REGION Network 13
   "V003 - Ventilador 3 Torres de enfriamiento Chillers"(Input_0 := "V003-TO",   // "FB_CTR_MOT"
                           Input_1 := "V003-CO",
                           Input_3 := ("DB90".Static_142 OR ("DB92".Static_12 AND NOT "DB90".Static_12)) AND NOT "DB86".Static_67 AND NOT "DB86".Static_68,
                           Input_6 := "UNO",
                           Input_7 := "DB90".Static_116,
                           Input_8 := "DB90".Static_12,
                           Output_0 => "V003-Marcha",
                           Output_2 => "DB32".Static_35,
                           Output_3 => "DB32".Static_36);
END_REGION

REGION Network 14
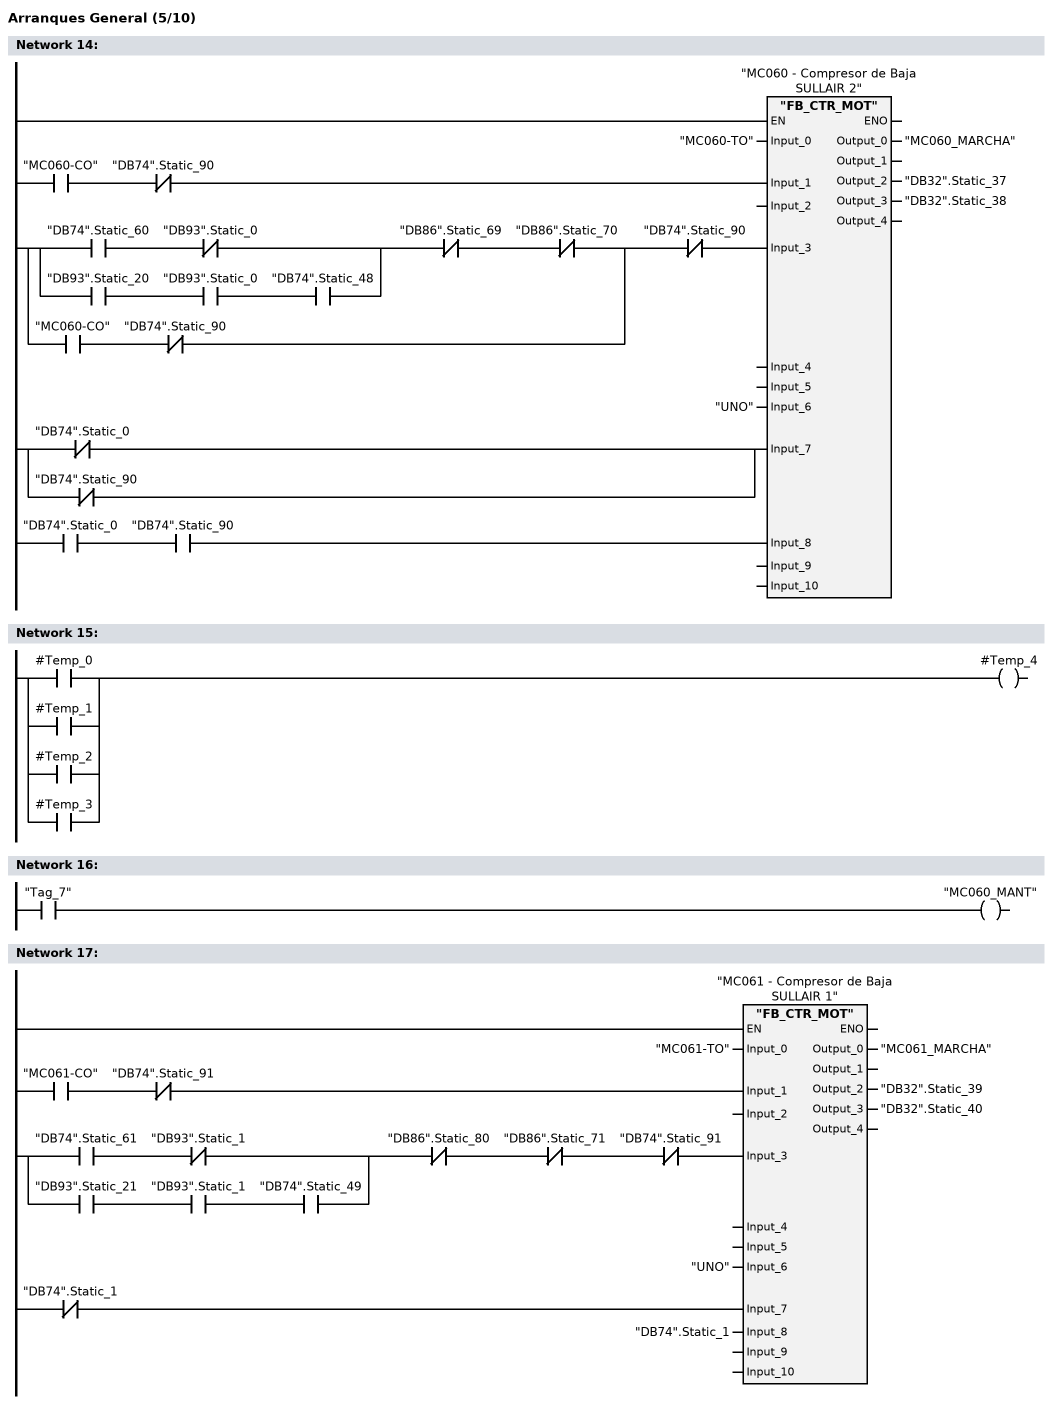
   "MC060 - Compresor de Baja SULLAIR 2"(Input_0 := "MC060-TO",   // "FB_CTR_MOT"
                           Input_1 := "MC060-CO" AND NOT "DB74".Static_90,
                           Input_3 := (((("DB74".Static_60 AND NOT "DB93".Static_0) OR ("DB93".Static_20 AND "DB93".Static_0 AND "DB74".Static_48)) AND NOT "DB86".Static_69 AND NOT "DB86".Static_70) OR ("MC060-CO" AND NOT "DB74".Static_90)) AND NOT "DB74".Static_90,
                           Input_6 := "UNO",
                           Input_7 := NOT "DB74".Static_0 OR NOT "DB74".Static_90,
                           Input_8 := "DB74".Static_0 AND "DB74".Static_90,
                           Output_0 => "MC060_MARCHA",
                           Output_2 => "DB32".Static_37,
                           Output_3 => "DB32".Static_38);
END_REGION

REGION Network 15
   RUNG wire#powerrail
      Contact( #Temp_0 )
      wire#w1
      Coil( #Temp_4 )
   END_RUNG
   RUNG wire#powerrail
      Contact( #Temp_1 )
   END_RUNG wire#w1
   RUNG wire#powerrail
      Contact( #Temp_2 )
   END_RUNG wire#w1
   RUNG wire#powerrail
      Contact( #Temp_3 )
   END_RUNG wire#w1
   // the same network as SCL:
   #Temp_4 := #Temp_0 OR #Temp_1 OR #Temp_2 OR #Temp_3;
END_REGION

REGION Network 16
   RUNG wire#powerrail
      Contact( "Tag_7" )
      Coil( "MC060_MANT" )
   END_RUNG
   // the same network as SCL:
   "MC060_MANT" := "Tag_7";
END_REGION

REGION Network 17
   RUNG wire#powerrail
      "MC061 - Compresor de Baja SULLAIR 1"(Input_0 := "MC061-TO", Input_2 :=, Input_4 :=, Input_5 :=, Input_6 := "UNO", Input_8 := "DB74".Static_1, Input_9 :=, Input_10 :=, Output_0 => "MC061_MARCHA", Output_1 =>, Output_2 => "DB32".Static_39, Output_3 => "DB32".Static_40, Output_4 =>, Input_1 := wire#w1, Input_3 := wire#w3, Input_7 := wire#w4)
   END_RUNG
   RUNG wire#powerrail
      Contact( "MC061-CO" )
      I_Contact( "DB74".Static_91 )
   END_RUNG wire#w1
   RUNG wire#powerrail
      Contact( "DB74".Static_61 )
      I_Contact( "DB93".Static_1 )
      wire#w2
      I_Contact( "DB86".Static_80 )
      I_Contact( "DB86".Static_71 )
      I_Contact( "DB74".Static_91 )
   END_RUNG wire#w3
   RUNG wire#powerrail
      Contact( "DB93".Static_21 )
      Contact( "DB93".Static_1 )
      Contact( "DB74".Static_49 )
   END_RUNG wire#w2
   RUNG wire#powerrail
      I_Contact( "DB74".Static_1 )
   END_RUNG wire#w4
   // the same network as SCL:
   "MC061 - Compresor de Baja SULLAIR 1"(Input_0 := "MC061-TO",   // "FB_CTR_MOT"
                           Input_1 := "MC061-CO" AND NOT "DB74".Static_91,
                           Input_3 := (("DB74".Static_61 AND NOT "DB93".Static_1) OR ("DB93".Static_21 AND "DB93".Static_1 AND "DB74".Static_49)) AND NOT "DB86".Static_80 AND NOT "DB86".Static_71 AND NOT "DB74".Static_91,
                           Input_6 := "UNO",
                           Input_7 := NOT "DB74".Static_1,
                           Input_8 := "DB74".Static_1,
                           Output_0 => "MC061_MARCHA",
                           Output_2 => "DB32".Static_39,
                           Output_3 => "DB32".Static_40);
END_REGION

REGION Network 18
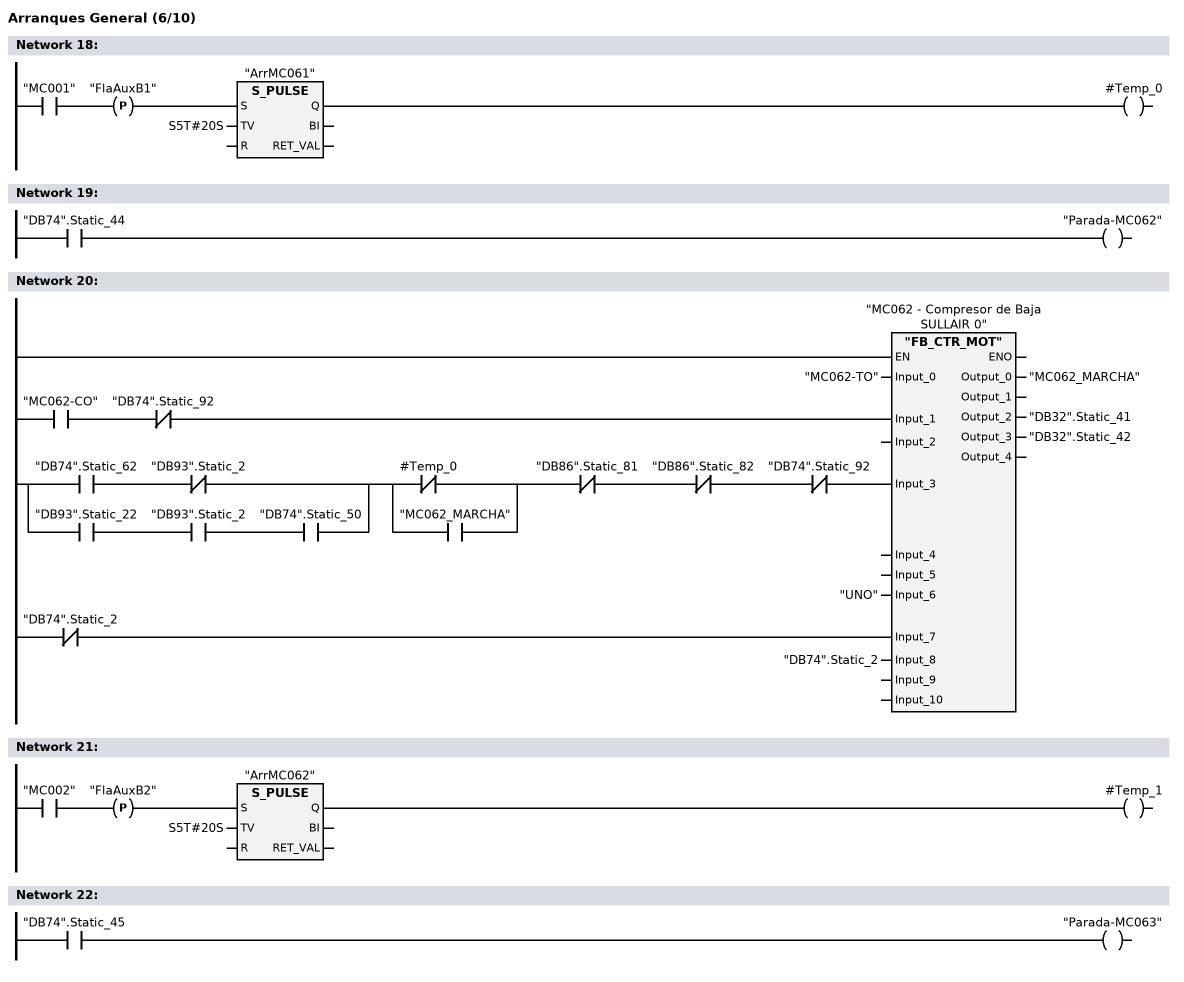
   RUNG wire#powerrail
      Contact( "MC001" )
      P_Trig( "FlaAuxB1" )
      S_PULSE(T_NO := "ArrMC061", TV := S5T#20S, R :=, BI =>, RET_VAL =>)
      Coil( #Temp_0 )
   END_RUNG
   // the same network as SCL:
   #_w1 := "MC001" AND NOT "FlaAuxB1";   // rising edge
   "FlaAuxB1" := "MC001";
   #_s5time1 := S_PULSE(T_NO := "ArrMC061", S := #_w1, TV := S5T#20S, Q => #_w2);
   #Temp_0 := #_w2;
END_REGION

REGION Network 19
   RUNG wire#powerrail
      Contact( "DB74".Static_44 )
      Coil( "Parada-MC062" )
   END_RUNG
   // the same network as SCL:
   "Parada-MC062" := "DB74".Static_44;
END_REGION

REGION Network 20
   RUNG wire#powerrail
      "MC062 - Compresor de Baja SULLAIR 0"(Input_0 := "MC062-TO", Input_2 :=, Input_4 :=, Input_5 :=, Input_6 := "UNO", Input_8 := "DB74".Static_2, Input_9 :=, Input_10 :=, Output_0 => "MC062_MARCHA", Output_1 =>, Output_2 => "DB32".Static_41, Output_3 => "DB32".Static_42, Output_4 =>, Input_1 := wire#w1, Input_3 := wire#w4, Input_7 := wire#w5)
   END_RUNG
   RUNG wire#powerrail
      Contact( "MC062-CO" )
      I_Contact( "DB74".Static_92 )
   END_RUNG wire#w1
   RUNG wire#powerrail
      Contact( "DB74".Static_62 )
      I_Contact( "DB93".Static_2 )
      wire#w2
      I_Contact( #Temp_0 )
      wire#w3
      I_Contact( "DB86".Static_81 )
      I_Contact( "DB86".Static_82 )
      I_Contact( "DB74".Static_92 )
   END_RUNG wire#w4
   RUNG wire#powerrail
      Contact( "DB93".Static_22 )
      Contact( "DB93".Static_2 )
      Contact( "DB74".Static_50 )
   END_RUNG wire#w2
   RUNG wire#w2
      Contact( "MC062_MARCHA" )
   END_RUNG wire#w3
   RUNG wire#powerrail
      I_Contact( "DB74".Static_2 )
   END_RUNG wire#w5
   // the same network as SCL:
   "MC062 - Compresor de Baja SULLAIR 0"(Input_0 := "MC062-TO",   // "FB_CTR_MOT"
                           Input_1 := "MC062-CO" AND NOT "DB74".Static_92,
                           Input_3 := (("DB74".Static_62 AND NOT "DB93".Static_2) OR ("DB93".Static_22 AND "DB93".Static_2 AND "DB74".Static_50)) AND (NOT #Temp_0 OR "MC062_MARCHA") AND NOT "DB86".Static_81 AND NOT "DB86".Static_82 AND NOT "DB74".Static_92,
                           Input_6 := "UNO",
                           Input_7 := NOT "DB74".Static_2,
                           Input_8 := "DB74".Static_2,
                           Output_0 => "MC062_MARCHA",
                           Output_2 => "DB32".Static_41,
                           Output_3 => "DB32".Static_42);
END_REGION

REGION Network 21
   RUNG wire#powerrail
      Contact( "MC002" )
      P_Trig( "FlaAuxB2" )
      S_PULSE(T_NO := "ArrMC062", TV := S5T#20S, R :=, BI =>, RET_VAL =>)
      Coil( #Temp_1 )
   END_RUNG
   // the same network as SCL:
   #_w1 := "MC002" AND NOT "FlaAuxB2";   // rising edge
   "FlaAuxB2" := "MC002";
   #_s5time1 := S_PULSE(T_NO := "ArrMC062", S := #_w1, TV := S5T#20S, Q => #_w2);
   #Temp_1 := #_w2;
END_REGION

REGION Network 22
   RUNG wire#powerrail
      Contact( "DB74".Static_45 )
      Coil( "Parada-MC063" )
   END_RUNG
   // the same network as SCL:
   "Parada-MC063" := "DB74".Static_45;
END_REGION

REGION Network 23
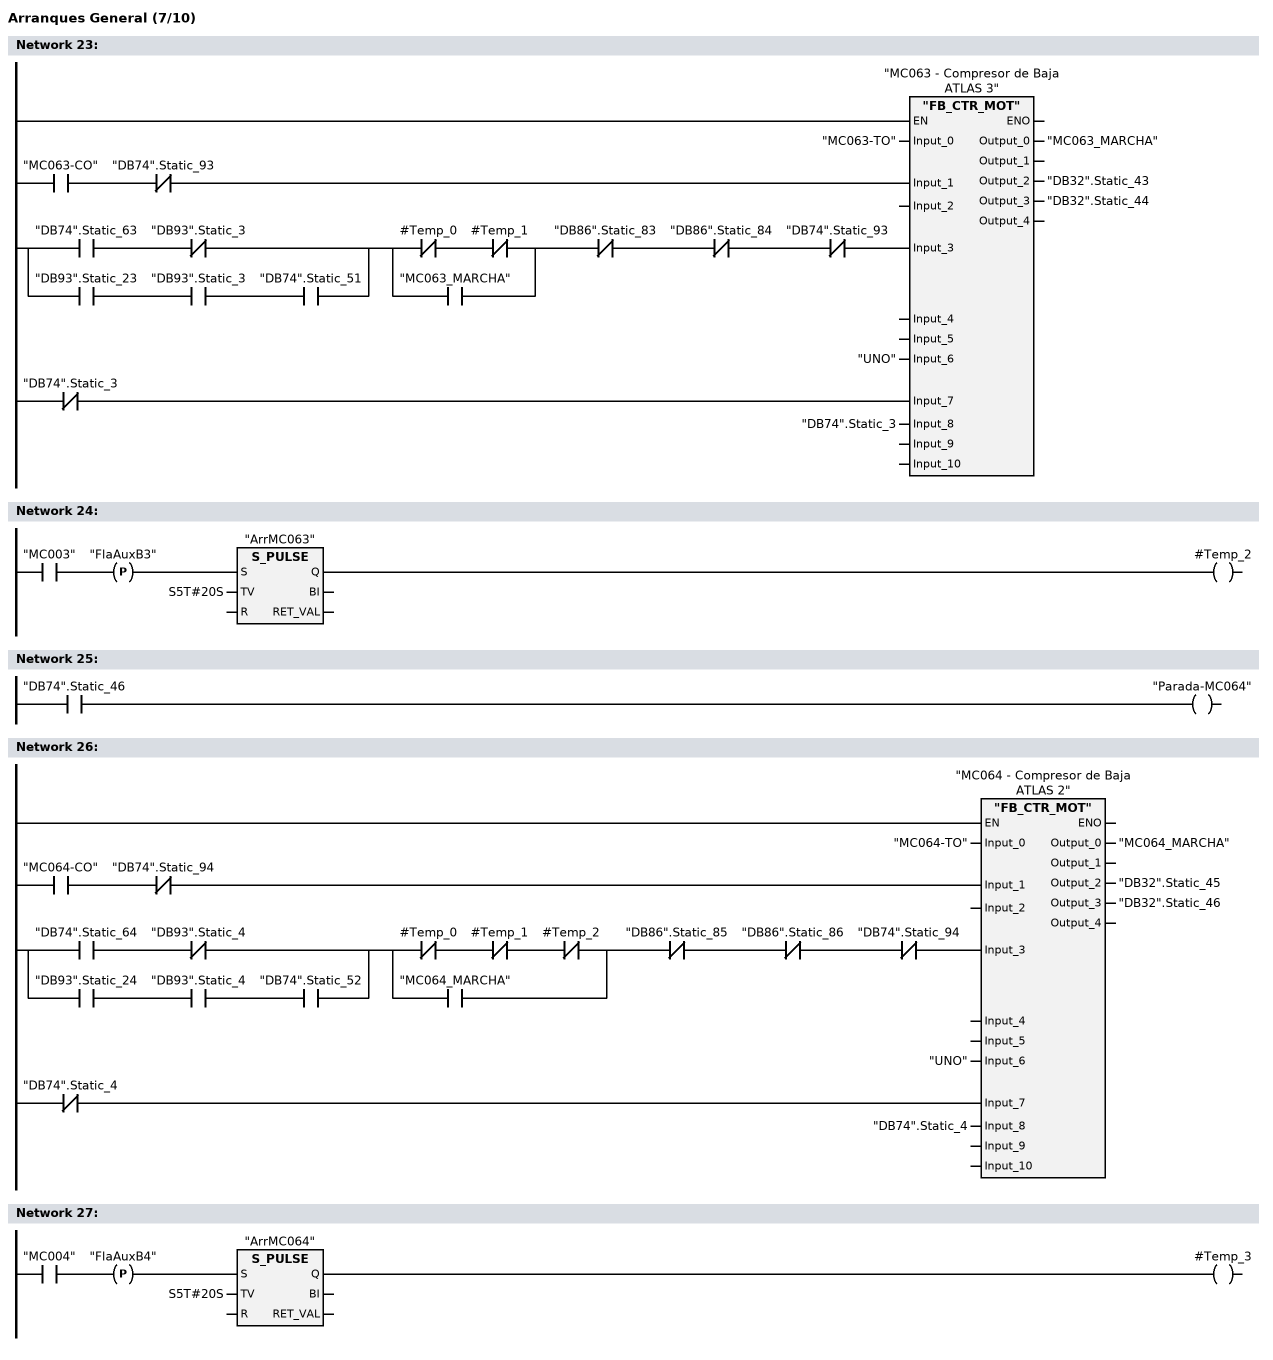
   RUNG wire#powerrail
      "MC063 - Compresor de Baja ATLAS 3"(Input_0 := "MC063-TO", Input_2 :=, Input_4 :=, Input_5 :=, Input_6 := "UNO", Input_8 := "DB74".Static_3, Input_9 :=, Input_10 :=, Output_0 => "MC063_MARCHA", Output_1 =>, Output_2 => "DB32".Static_43, Output_3 => "DB32".Static_44, Output_4 =>, Input_1 := wire#w1, Input_3 := wire#w4, Input_7 := wire#w5)
   END_RUNG
   RUNG wire#powerrail
      Contact( "MC063-CO" )
      I_Contact( "DB74".Static_93 )
   END_RUNG wire#w1
   RUNG wire#powerrail
      Contact( "DB74".Static_63 )
      I_Contact( "DB93".Static_3 )
      wire#w2
      I_Contact( #Temp_0 )
      I_Contact( #Temp_1 )
      wire#w3
      I_Contact( "DB86".Static_83 )
      I_Contact( "DB86".Static_84 )
      I_Contact( "DB74".Static_93 )
   END_RUNG wire#w4
   RUNG wire#powerrail
      Contact( "DB93".Static_23 )
      Contact( "DB93".Static_3 )
      Contact( "DB74".Static_51 )
   END_RUNG wire#w2
   RUNG wire#w2
      Contact( "MC063_MARCHA" )
   END_RUNG wire#w3
   RUNG wire#powerrail
      I_Contact( "DB74".Static_3 )
   END_RUNG wire#w5
   // the same network as SCL:
   "MC063 - Compresor de Baja ATLAS 3"(Input_0 := "MC063-TO",   // "FB_CTR_MOT"
                           Input_1 := "MC063-CO" AND NOT "DB74".Static_93,
                           Input_3 := (("DB74".Static_63 AND NOT "DB93".Static_3) OR ("DB93".Static_23 AND "DB93".Static_3 AND "DB74".Static_51)) AND ((NOT #Temp_0 AND NOT #Temp_1) OR "MC063_MARCHA") AND NOT "DB86".Static_83 AND NOT "DB86".Static_84 AND NOT "DB74".Static_93,
                           Input_6 := "UNO",
                           Input_7 := NOT "DB74".Static_3,
                           Input_8 := "DB74".Static_3,
                           Output_0 => "MC063_MARCHA",
                           Output_2 => "DB32".Static_43,
                           Output_3 => "DB32".Static_44);
END_REGION

REGION Network 24
   RUNG wire#powerrail
      Contact( "MC003" )
      P_Trig( "FlaAuxB3" )
      S_PULSE(T_NO := "ArrMC063", TV := S5T#20S, R :=, BI =>, RET_VAL =>)
      Coil( #Temp_2 )
   END_RUNG
   // the same network as SCL:
   #_w1 := "MC003" AND NOT "FlaAuxB3";   // rising edge
   "FlaAuxB3" := "MC003";
   #_s5time1 := S_PULSE(T_NO := "ArrMC063", S := #_w1, TV := S5T#20S, Q => #_w2);
   #Temp_2 := #_w2;
END_REGION

REGION Network 25
   RUNG wire#powerrail
      Contact( "DB74".Static_46 )
      Coil( "Parada-MC064" )
   END_RUNG
   // the same network as SCL:
   "Parada-MC064" := "DB74".Static_46;
END_REGION

REGION Network 26
   RUNG wire#powerrail
      "MC064 - Compresor de Baja ATLAS 2"(Input_0 := "MC064-TO", Input_2 :=, Input_4 :=, Input_5 :=, Input_6 := "UNO", Input_8 := "DB74".Static_4, Input_9 :=, Input_10 :=, Output_0 => "MC064_MARCHA", Output_1 =>, Output_2 => "DB32".Static_45, Output_3 => "DB32".Static_46, Output_4 =>, Input_1 := wire#w1, Input_3 := wire#w4, Input_7 := wire#w5)
   END_RUNG
   RUNG wire#powerrail
      Contact( "MC064-CO" )
      I_Contact( "DB74".Static_94 )
   END_RUNG wire#w1
   RUNG wire#powerrail
      Contact( "DB74".Static_64 )
      I_Contact( "DB93".Static_4 )
      wire#w2
      I_Contact( #Temp_0 )
      I_Contact( #Temp_1 )
      I_Contact( #Temp_2 )
      wire#w3
      I_Contact( "DB86".Static_85 )
      I_Contact( "DB86".Static_86 )
      I_Contact( "DB74".Static_94 )
   END_RUNG wire#w4
   RUNG wire#powerrail
      Contact( "DB93".Static_24 )
      Contact( "DB93".Static_4 )
      Contact( "DB74".Static_52 )
   END_RUNG wire#w2
   RUNG wire#w2
      Contact( "MC064_MARCHA" )
   END_RUNG wire#w3
   RUNG wire#powerrail
      I_Contact( "DB74".Static_4 )
   END_RUNG wire#w5
   // the same network as SCL:
   "MC064 - Compresor de Baja ATLAS 2"(Input_0 := "MC064-TO",   // "FB_CTR_MOT"
                           Input_1 := "MC064-CO" AND NOT "DB74".Static_94,
                           Input_3 := (("DB74".Static_64 AND NOT "DB93".Static_4) OR ("DB93".Static_24 AND "DB93".Static_4 AND "DB74".Static_52)) AND ((NOT #Temp_0 AND NOT #Temp_1 AND NOT #Temp_2) OR "MC064_MARCHA") AND NOT "DB86".Static_85 AND NOT "DB86".Static_86 AND NOT "DB74".Static_94,
                           Input_6 := "UNO",
                           Input_7 := NOT "DB74".Static_4,
                           Input_8 := "DB74".Static_4,
                           Output_0 => "MC064_MARCHA",
                           Output_2 => "DB32".Static_45,
                           Output_3 => "DB32".Static_46);
END_REGION

REGION Network 27
   RUNG wire#powerrail
      Contact( "MC004" )
      P_Trig( "FlaAuxB4" )
      S_PULSE(T_NO := "ArrMC064", TV := S5T#20S, R :=, BI =>, RET_VAL =>)
      Coil( #Temp_3 )
   END_RUNG
   // the same network as SCL:
   #_w1 := "MC004" AND NOT "FlaAuxB4";   // rising edge
   "FlaAuxB4" := "MC004";
   #_s5time1 := S_PULSE(T_NO := "ArrMC064", S := #_w1, TV := S5T#20S, Q => #_w2);
   #Temp_3 := #_w2;
END_REGION

REGION Network 28
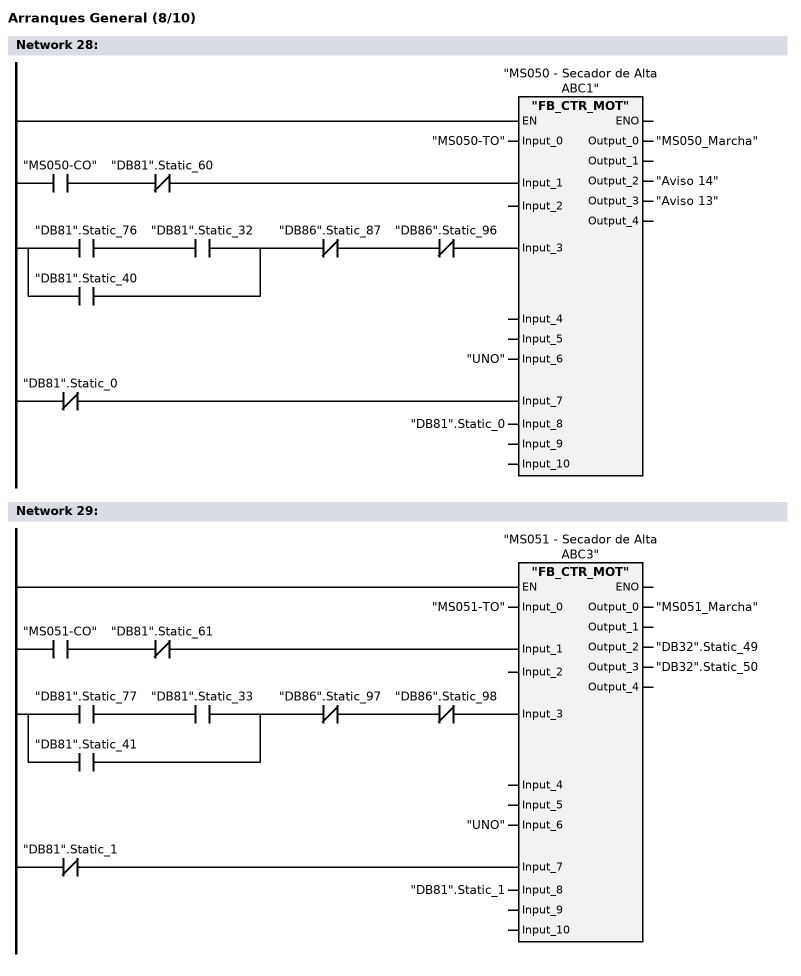
   "MS050 - Secador de Alta  ABC1"(Input_0 := "MS050-TO",   // "FB_CTR_MOT"
                           Input_1 := "MS050-CO" AND NOT "DB81".Static_60,
                           Input_3 := ("DB81".Static_40 OR ("DB81".Static_76 AND "DB81".Static_32)) AND NOT "DB86".Static_87 AND NOT "DB86".Static_96,
                           Input_6 := "UNO",
                           Input_7 := NOT "DB81".Static_0,
                           Input_8 := "DB81".Static_0,
                           Output_0 => "MS050_Marcha",
                           Output_2 => "Aviso 14",
                           Output_3 => "Aviso 13");
END_REGION

REGION Network 29
   "MS051 - Secador de Alta  ABC3"(Input_0 := "MS051-TO",   // "FB_CTR_MOT"
                           Input_1 := "MS051-CO" AND NOT "DB81".Static_61,
                           Input_3 := ("DB81".Static_41 OR ("DB81".Static_77 AND "DB81".Static_33)) AND NOT "DB86".Static_97 AND NOT "DB86".Static_98,
                           Input_6 := "UNO",
                           Input_7 := NOT "DB81".Static_1,
                           Input_8 := "DB81".Static_1,
                           Output_0 => "MS051_Marcha",
                           Output_2 => "DB32".Static_49,
                           Output_3 => "DB32".Static_50);
END_REGION

REGION Network 30
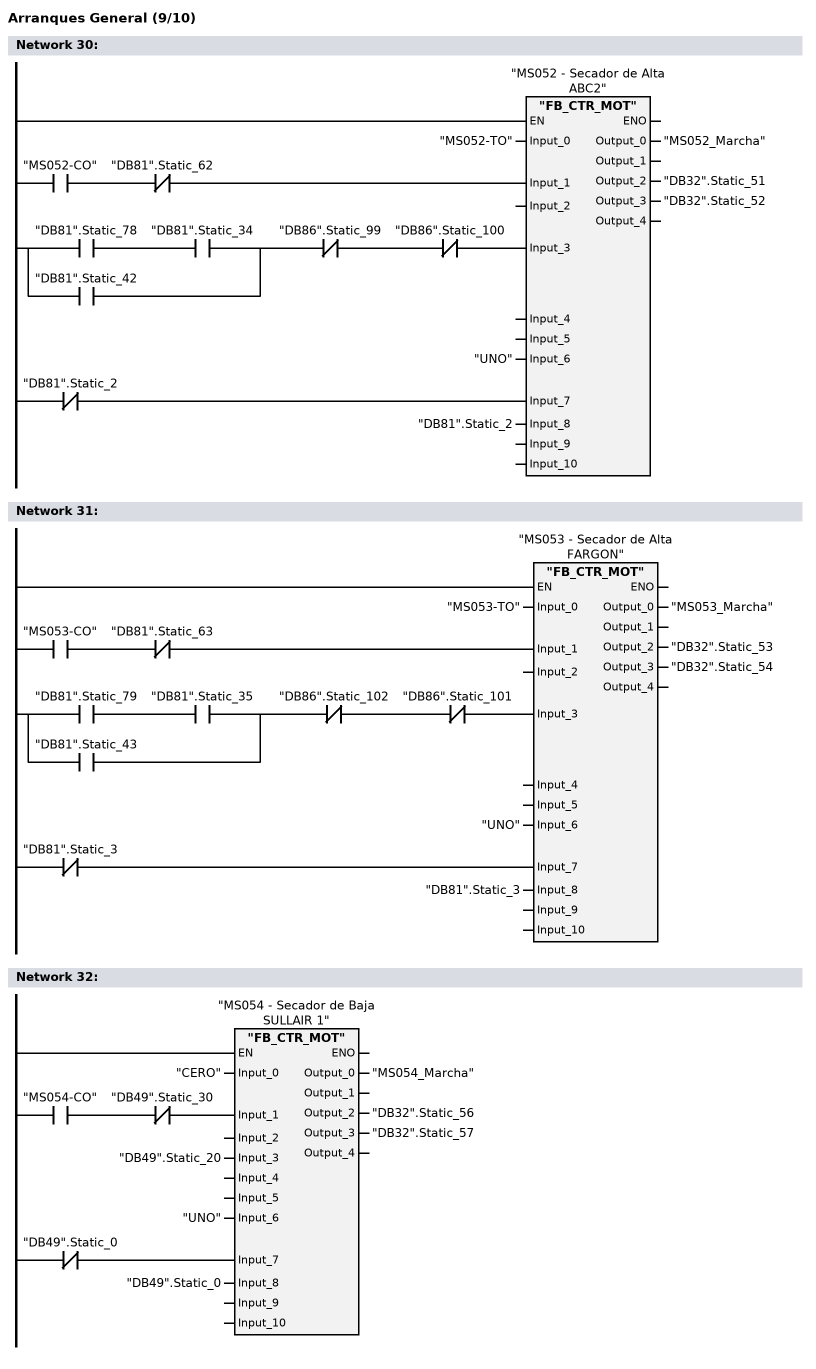
   "MS052 - Secador de Alta  ABC2"(Input_0 := "MS052-TO",   // "FB_CTR_MOT"
                           Input_1 := "MS052-CO" AND NOT "DB81".Static_62,
                           Input_3 := ("DB81".Static_42 OR ("DB81".Static_78 AND "DB81".Static_34)) AND NOT "DB86".Static_99 AND NOT "DB86".Static_100,
                           Input_6 := "UNO",
                           Input_7 := NOT "DB81".Static_2,
                           Input_8 := "DB81".Static_2,
                           Output_0 => "MS052_Marcha",
                           Output_2 => "DB32".Static_51,
                           Output_3 => "DB32".Static_52);
END_REGION

REGION Network 31
   "MS053 - Secador de Alta  FARGON"(Input_0 := "MS053-TO",   // "FB_CTR_MOT"
                           Input_1 := "MS053-CO" AND NOT "DB81".Static_63,
                           Input_3 := ("DB81".Static_43 OR ("DB81".Static_79 AND "DB81".Static_35)) AND NOT "DB86".Static_102 AND NOT "DB86".Static_101,
                           Input_6 := "UNO",
                           Input_7 := NOT "DB81".Static_3,
                           Input_8 := "DB81".Static_3,
                           Output_0 => "MS053_Marcha",
                           Output_2 => "DB32".Static_53,
                           Output_3 => "DB32".Static_54);
END_REGION

REGION Network 32
   RUNG wire#powerrail
      "MS054 - Secador de Baja SULLAIR 1"(Input_0 := "CERO", Input_2 :=, Input_3 := "DB49".Static_20, Input_4 :=, Input_5 :=, Input_6 := "UNO", Input_8 := "DB49".Static_0, Input_9 :=, Input_10 :=, Output_0 => "MS054_Marcha", Output_1 =>, Output_2 => "DB32".Static_56, Output_3 => "DB32".Static_57, Output_4 =>, Input_1 := wire#w1, Input_7 := wire#w2)
   END_RUNG
   RUNG wire#powerrail
      Contact( "MS054-CO" )
      I_Contact( "DB49".Static_30 )
   END_RUNG wire#w1
   RUNG wire#powerrail
      I_Contact( "DB49".Static_0 )
   END_RUNG wire#w2
   // the same network as SCL:
   "MS054 - Secador de Baja SULLAIR 1"(Input_0 := "CERO",   // "FB_CTR_MOT"
                           Input_1 := "MS054-CO" AND NOT "DB49".Static_30,
                           Input_3 := "DB49".Static_20,
                           Input_6 := "UNO",
                           Input_7 := NOT "DB49".Static_0,
                           Input_8 := "DB49".Static_0,
                           Output_0 => "MS054_Marcha",
                           Output_2 => "DB32".Static_56,
                           Output_3 => "DB32".Static_57);
END_REGION

REGION Network 33
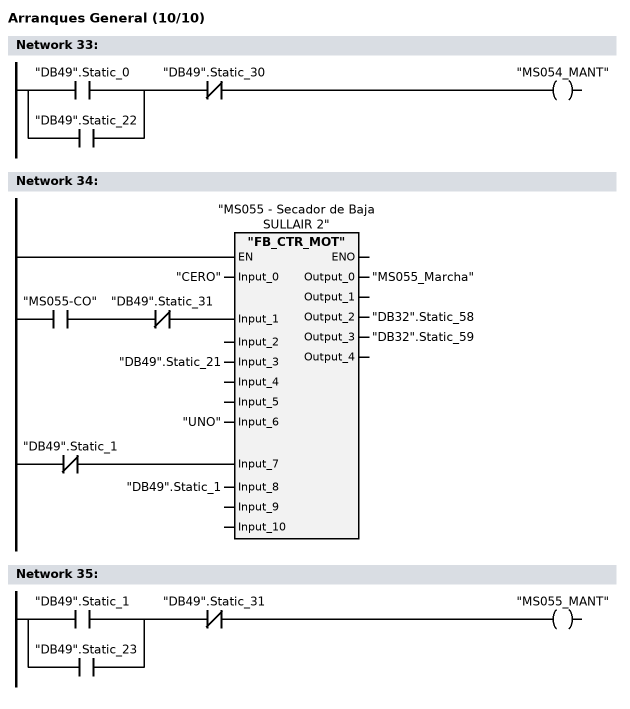
   RUNG wire#powerrail
      Contact( "DB49".Static_0 )
      wire#w1
      I_Contact( "DB49".Static_30 )
      Coil( "MS054_MANT" )
   END_RUNG
   RUNG wire#powerrail
      Contact( "DB49".Static_22 )
   END_RUNG wire#w1
   // the same network as SCL:
   "MS054_MANT" := ("DB49".Static_0 OR "DB49".Static_22) AND NOT "DB49".Static_30;
END_REGION

REGION Network 34
   RUNG wire#powerrail
      "MS055 - Secador de Baja SULLAIR 2"(Input_0 := "CERO", Input_2 :=, Input_3 := "DB49".Static_21, Input_4 :=, Input_5 :=, Input_6 := "UNO", Input_8 := "DB49".Static_1, Input_9 :=, Input_10 :=, Output_0 => "MS055_Marcha", Output_1 =>, Output_2 => "DB32".Static_58, Output_3 => "DB32".Static_59, Output_4 =>, Input_1 := wire#w1, Input_7 := wire#w2)
   END_RUNG
   RUNG wire#powerrail
      Contact( "MS055-CO" )
      I_Contact( "DB49".Static_31 )
   END_RUNG wire#w1
   RUNG wire#powerrail
      I_Contact( "DB49".Static_1 )
   END_RUNG wire#w2
   // the same network as SCL:
   "MS055 - Secador de Baja SULLAIR 2"(Input_0 := "CERO",   // "FB_CTR_MOT"
                           Input_1 := "MS055-CO" AND NOT "DB49".Static_31,
                           Input_3 := "DB49".Static_21,
                           Input_6 := "UNO",
                           Input_7 := NOT "DB49".Static_1,
                           Input_8 := "DB49".Static_1,
                           Output_0 => "MS055_Marcha",
                           Output_2 => "DB32".Static_58,
                           Output_3 => "DB32".Static_59);
END_REGION

REGION Network 35
   RUNG wire#powerrail
      Contact( "DB49".Static_1 )
      wire#w1
      I_Contact( "DB49".Static_31 )
      Coil( "MS055_MANT" )
   END_RUNG
   RUNG wire#powerrail
      Contact( "DB49".Static_23 )
   END_RUNG wire#w1
   // the same network as SCL:
   "MS055_MANT" := ("DB49".Static_1 OR "DB49".Static_23) AND NOT "DB49".Static_31;
END_REGION
END_FUNCTION

FUNCTION "FC51" : Void   // FC51, LAD
{ S7_Optimized_Access := 'FALSE' }
VERSION : 0.1
   VAR_TEMP   // added for the SCL form of the ladder/FBD networks
      _w1 : Bool;
      _s5time1 : S5Time;
      _s5time2 : S5Time;
   END_VAR
BEGIN

REGION Network 1
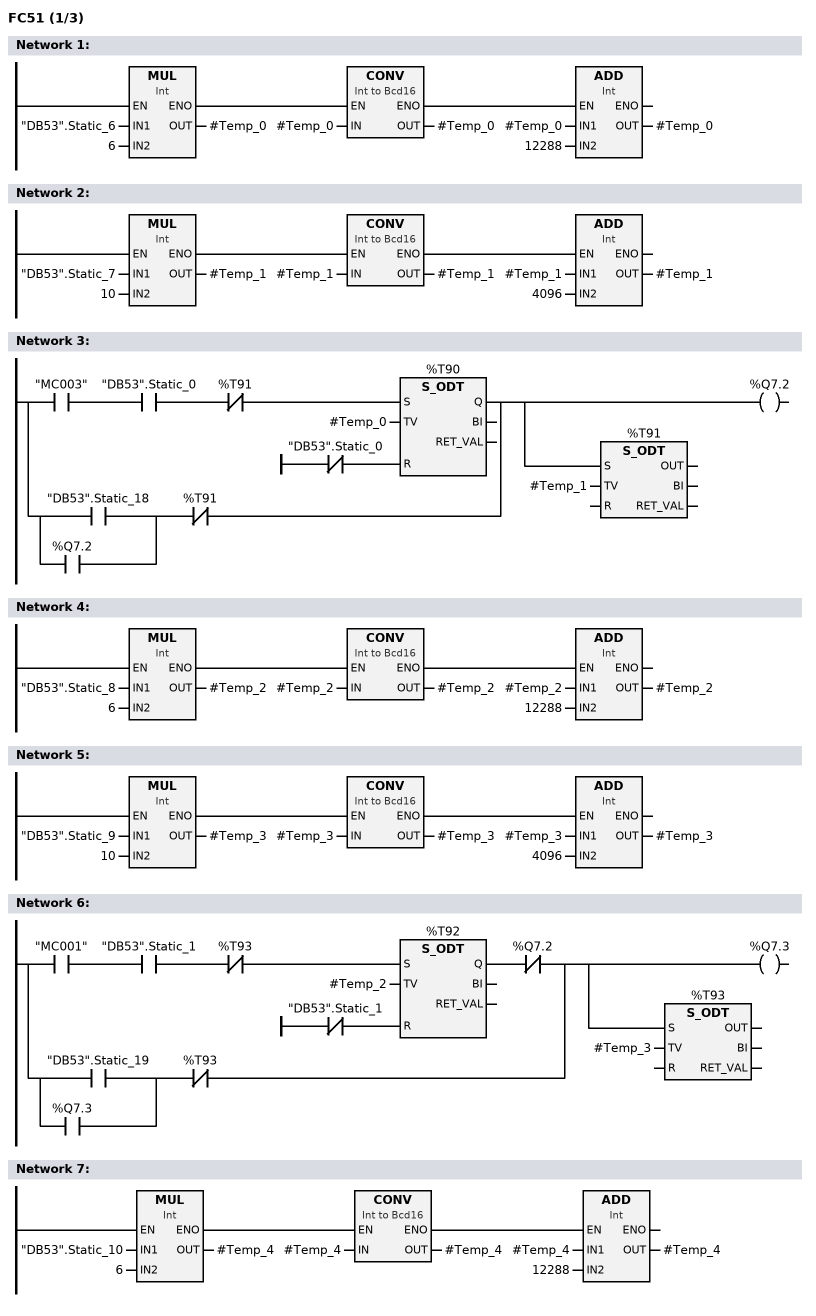
   RUNG wire#powerrail
      { S7_Templates := "SrcType := Int"; S7_GenerateENO := "TRUE" } Mul(in1 := "DB53".Static_6, in2 := 6, out => #Temp_0)
      { S7_Templates := "[SrcType := Int, DestType := Bcd16]"; S7_GenerateENO := "TRUE" } Convert(in := #Temp_0, out => #Temp_0)
      { S7_Templates := "SrcType := Int"; S7_GenerateENO := "TRUE" } Add(in1 := #Temp_0, in2 := 12288, out => #Temp_0)
   END_RUNG
   // the same network as SCL:
   // ENO of a box is taken as its EN; it also drops when the box reports an error
   #Temp_0 := "DB53".Static_6 * 6;
   #Temp_0 := INT_TO_BCD16(#Temp_0);
   #Temp_0 := #Temp_0 + 12288;
END_REGION

REGION Network 2
   RUNG wire#powerrail
      { S7_Templates := "SrcType := Int"; S7_GenerateENO := "TRUE" } Mul(in1 := "DB53".Static_7, in2 := 10, out => #Temp_1)
      { S7_Templates := "[SrcType := Int, DestType := Bcd16]"; S7_GenerateENO := "TRUE" } Convert(in := #Temp_1, out => #Temp_1)
      { S7_Templates := "SrcType := Int"; S7_GenerateENO := "TRUE" } Add(in1 := #Temp_1, in2 := 4096, out => #Temp_1)
   END_RUNG
   // the same network as SCL:
   // ENO of a box is taken as its EN; it also drops when the box reports an error
   #Temp_1 := "DB53".Static_7 * 10;
   #Temp_1 := INT_TO_BCD16(#Temp_1);
   #Temp_1 := #Temp_1 + 4096;
END_REGION

REGION Network 3
   RUNG wire#powerrail
      Contact( "MC003" )
      Contact( "DB53".Static_0 )
      I_Contact( %T91 )
      S_ODT(T_NO := %T90, TV := #Temp_0, R := wire#w1, BI =>, RET_VAL =>)
      wire#w2
      Coil( %Q7.2 )
   END_RUNG
   RUNG wire#powerrail
      I_Contact( "DB53".Static_0 )
   END_RUNG wire#w1
   RUNG wire#powerrail
      Contact( "DB53".Static_18 )
      wire#w3
      I_Contact( %T91 )
   END_RUNG wire#w2
   RUNG wire#powerrail
      Contact( %Q7.2 )
   END_RUNG wire#w3
   RUNG wire#w2
      S_ODT(T_NO := %T91, TV := #Temp_1, R :=, BI =>, RET_VAL =>)
   END_RUNG
   // the same network as SCL:
   #_s5time1 := S_ODT(T_NO := %T90,
                      TV := #Temp_0,
                      S := "MC003" AND "DB53".Static_0 AND NOT %T91,
                      R := NOT "DB53".Static_0,
                      Q => #_w1);
   %Q7.2 := #_w1 OR (("DB53".Static_18 OR %Q7.2) AND NOT %T91);
   #_s5time2 := S_ODT(T_NO := %T91, TV := #Temp_1, S := %Q7.2);
END_REGION

REGION Network 4
   RUNG wire#powerrail
      { S7_Templates := "SrcType := Int"; S7_GenerateENO := "TRUE" } Mul(in1 := "DB53".Static_8, in2 := 6, out => #Temp_2)
      { S7_Templates := "[SrcType := Int, DestType := Bcd16]"; S7_GenerateENO := "TRUE" } Convert(in := #Temp_2, out => #Temp_2)
      { S7_Templates := "SrcType := Int"; S7_GenerateENO := "TRUE" } Add(in1 := #Temp_2, in2 := 12288, out => #Temp_2)
   END_RUNG
   // the same network as SCL:
   // ENO of a box is taken as its EN; it also drops when the box reports an error
   #Temp_2 := "DB53".Static_8 * 6;
   #Temp_2 := INT_TO_BCD16(#Temp_2);
   #Temp_2 := #Temp_2 + 12288;
END_REGION

REGION Network 5
   RUNG wire#powerrail
      { S7_Templates := "SrcType := Int"; S7_GenerateENO := "TRUE" } Mul(in1 := "DB53".Static_9, in2 := 10, out => #Temp_3)
      { S7_Templates := "[SrcType := Int, DestType := Bcd16]"; S7_GenerateENO := "TRUE" } Convert(in := #Temp_3, out => #Temp_3)
      { S7_Templates := "SrcType := Int"; S7_GenerateENO := "TRUE" } Add(in1 := #Temp_3, in2 := 4096, out => #Temp_3)
   END_RUNG
   // the same network as SCL:
   // ENO of a box is taken as its EN; it also drops when the box reports an error
   #Temp_3 := "DB53".Static_9 * 10;
   #Temp_3 := INT_TO_BCD16(#Temp_3);
   #Temp_3 := #Temp_3 + 4096;
END_REGION

REGION Network 6
   RUNG wire#powerrail
      Contact( "MC001" )
      Contact( "DB53".Static_1 )
      I_Contact( %T93 )
      S_ODT(T_NO := %T92, TV := #Temp_2, R := wire#w1, BI =>, RET_VAL =>)
      I_Contact( %Q7.2 )
      wire#w2
      Coil( %Q7.3 )
   END_RUNG
   RUNG wire#powerrail
      I_Contact( "DB53".Static_1 )
   END_RUNG wire#w1
   RUNG wire#powerrail
      Contact( "DB53".Static_19 )
      wire#w3
      I_Contact( %T93 )
   END_RUNG wire#w2
   RUNG wire#powerrail
      Contact( %Q7.3 )
   END_RUNG wire#w3
   RUNG wire#w2
      S_ODT(T_NO := %T93, TV := #Temp_3, R :=, BI =>, RET_VAL =>)
   END_RUNG
   // the same network as SCL:
   #_s5time1 := S_ODT(T_NO := %T92,
                      TV := #Temp_2,
                      S := "MC001" AND "DB53".Static_1 AND NOT %T93,
                      R := NOT "DB53".Static_1,
                      Q => #_w1);
   %Q7.3 := (#_w1 AND NOT %Q7.2) OR (("DB53".Static_19 OR %Q7.3) AND NOT %T93);
   #_s5time2 := S_ODT(T_NO := %T93, TV := #Temp_3, S := %Q7.3);
END_REGION

REGION Network 7
   RUNG wire#powerrail
      { S7_Templates := "SrcType := Int"; S7_GenerateENO := "TRUE" } Mul(in1 := "DB53".Static_10, in2 := 6, out => #Temp_4)
      { S7_Templates := "[SrcType := Int, DestType := Bcd16]"; S7_GenerateENO := "TRUE" } Convert(in := #Temp_4, out => #Temp_4)
      { S7_Templates := "SrcType := Int"; S7_GenerateENO := "TRUE" } Add(in1 := #Temp_4, in2 := 12288, out => #Temp_4)
   END_RUNG
   // the same network as SCL:
   // ENO of a box is taken as its EN; it also drops when the box reports an error
   #Temp_4 := "DB53".Static_10 * 6;
   #Temp_4 := INT_TO_BCD16(#Temp_4);
   #Temp_4 := #Temp_4 + 12288;
END_REGION

REGION Network 8
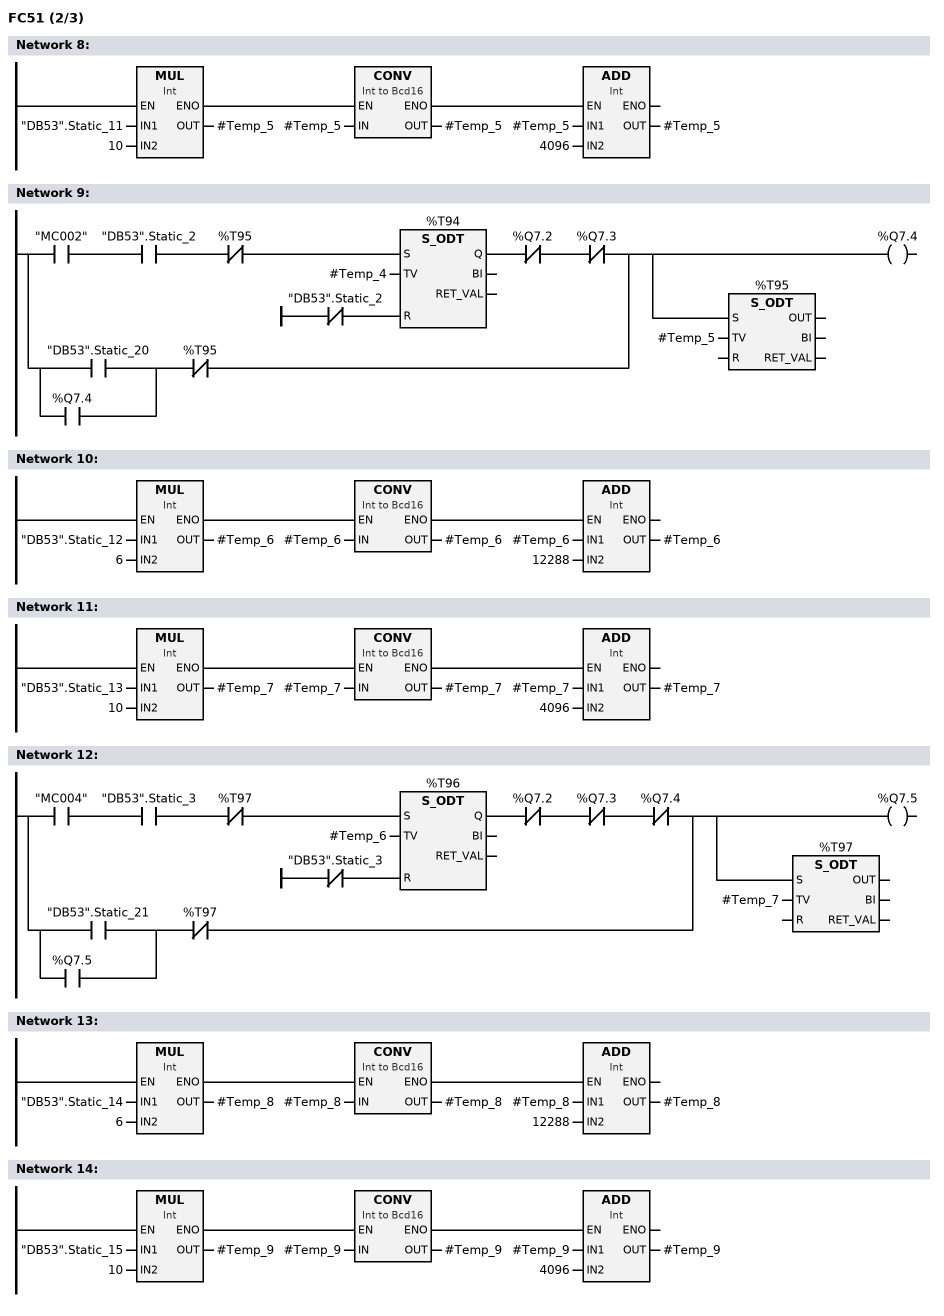
   RUNG wire#powerrail
      { S7_Templates := "SrcType := Int"; S7_GenerateENO := "TRUE" } Mul(in1 := "DB53".Static_11, in2 := 10, out => #Temp_5)
      { S7_Templates := "[SrcType := Int, DestType := Bcd16]"; S7_GenerateENO := "TRUE" } Convert(in := #Temp_5, out => #Temp_5)
      { S7_Templates := "SrcType := Int"; S7_GenerateENO := "TRUE" } Add(in1 := #Temp_5, in2 := 4096, out => #Temp_5)
   END_RUNG
   // the same network as SCL:
   // ENO of a box is taken as its EN; it also drops when the box reports an error
   #Temp_5 := "DB53".Static_11 * 10;
   #Temp_5 := INT_TO_BCD16(#Temp_5);
   #Temp_5 := #Temp_5 + 4096;
END_REGION

REGION Network 9
   RUNG wire#powerrail
      Contact( "MC002" )
      Contact( "DB53".Static_2 )
      I_Contact( %T95 )
      S_ODT(T_NO := %T94, TV := #Temp_4, R := wire#w1, BI =>, RET_VAL =>)
      I_Contact( %Q7.2 )
      I_Contact( %Q7.3 )
      wire#w2
      Coil( %Q7.4 )
   END_RUNG
   RUNG wire#powerrail
      I_Contact( "DB53".Static_2 )
   END_RUNG wire#w1
   RUNG wire#powerrail
      Contact( "DB53".Static_20 )
      wire#w3
      I_Contact( %T95 )
   END_RUNG wire#w2
   RUNG wire#powerrail
      Contact( %Q7.4 )
   END_RUNG wire#w3
   RUNG wire#w2
      S_ODT(T_NO := %T95, TV := #Temp_5, R :=, BI =>, RET_VAL =>)
   END_RUNG
   // the same network as SCL:
   #_s5time1 := S_ODT(T_NO := %T94,
                      TV := #Temp_4,
                      S := "MC002" AND "DB53".Static_2 AND NOT %T95,
                      R := NOT "DB53".Static_2,
                      Q => #_w1);
   %Q7.4 := (#_w1 AND NOT %Q7.2 AND NOT %Q7.3) OR (("DB53".Static_20 OR %Q7.4) AND NOT %T95);
   #_s5time2 := S_ODT(T_NO := %T95, TV := #Temp_5, S := %Q7.4);
END_REGION

REGION Network 10
   RUNG wire#powerrail
      { S7_Templates := "SrcType := Int"; S7_GenerateENO := "TRUE" } Mul(in1 := "DB53".Static_12, in2 := 6, out => #Temp_6)
      { S7_Templates := "[SrcType := Int, DestType := Bcd16]"; S7_GenerateENO := "TRUE" } Convert(in := #Temp_6, out => #Temp_6)
      { S7_Templates := "SrcType := Int"; S7_GenerateENO := "TRUE" } Add(in1 := #Temp_6, in2 := 12288, out => #Temp_6)
   END_RUNG
   // the same network as SCL:
   // ENO of a box is taken as its EN; it also drops when the box reports an error
   #Temp_6 := "DB53".Static_12 * 6;
   #Temp_6 := INT_TO_BCD16(#Temp_6);
   #Temp_6 := #Temp_6 + 12288;
END_REGION

REGION Network 11
   RUNG wire#powerrail
      { S7_Templates := "SrcType := Int"; S7_GenerateENO := "TRUE" } Mul(in1 := "DB53".Static_13, in2 := 10, out => #Temp_7)
      { S7_Templates := "[SrcType := Int, DestType := Bcd16]"; S7_GenerateENO := "TRUE" } Convert(in := #Temp_7, out => #Temp_7)
      { S7_Templates := "SrcType := Int"; S7_GenerateENO := "TRUE" } Add(in1 := #Temp_7, in2 := 4096, out => #Temp_7)
   END_RUNG
   // the same network as SCL:
   // ENO of a box is taken as its EN; it also drops when the box reports an error
   #Temp_7 := "DB53".Static_13 * 10;
   #Temp_7 := INT_TO_BCD16(#Temp_7);
   #Temp_7 := #Temp_7 + 4096;
END_REGION

REGION Network 12
   RUNG wire#powerrail
      Contact( "MC004" )
      Contact( "DB53".Static_3 )
      I_Contact( %T97 )
      S_ODT(T_NO := %T96, TV := #Temp_6, R := wire#w1, BI =>, RET_VAL =>)
      I_Contact( %Q7.2 )
      I_Contact( %Q7.3 )
      I_Contact( %Q7.4 )
      wire#w2
      Coil( %Q7.5 )
   END_RUNG
   RUNG wire#powerrail
      I_Contact( "DB53".Static_3 )
   END_RUNG wire#w1
   RUNG wire#powerrail
      Contact( "DB53".Static_21 )
      wire#w3
      I_Contact( %T97 )
   END_RUNG wire#w2
   RUNG wire#powerrail
      Contact( %Q7.5 )
   END_RUNG wire#w3
   RUNG wire#w2
      S_ODT(T_NO := %T97, TV := #Temp_7, R :=, BI =>, RET_VAL =>)
   END_RUNG
   // the same network as SCL:
   #_s5time1 := S_ODT(T_NO := %T96,
                      TV := #Temp_6,
                      S := "MC004" AND "DB53".Static_3 AND NOT %T97,
                      R := NOT "DB53".Static_3,
                      Q => #_w1);
   %Q7.5 := (#_w1 AND NOT %Q7.2 AND NOT %Q7.3 AND NOT %Q7.4) OR (("DB53".Static_21 OR %Q7.5) AND NOT %T97);
   #_s5time2 := S_ODT(T_NO := %T97, TV := #Temp_7, S := %Q7.5);
END_REGION

REGION Network 13
   RUNG wire#powerrail
      { S7_Templates := "SrcType := Int"; S7_GenerateENO := "TRUE" } Mul(in1 := "DB53".Static_14, in2 := 6, out => #Temp_8)
      { S7_Templates := "[SrcType := Int, DestType := Bcd16]"; S7_GenerateENO := "TRUE" } Convert(in := #Temp_8, out => #Temp_8)
      { S7_Templates := "SrcType := Int"; S7_GenerateENO := "TRUE" } Add(in1 := #Temp_8, in2 := 12288, out => #Temp_8)
   END_RUNG
   // the same network as SCL:
   // ENO of a box is taken as its EN; it also drops when the box reports an error
   #Temp_8 := "DB53".Static_14 * 6;
   #Temp_8 := INT_TO_BCD16(#Temp_8);
   #Temp_8 := #Temp_8 + 12288;
END_REGION

REGION Network 14
   RUNG wire#powerrail
      { S7_Templates := "SrcType := Int"; S7_GenerateENO := "TRUE" } Mul(in1 := "DB53".Static_15, in2 := 10, out => #Temp_9)
      { S7_Templates := "[SrcType := Int, DestType := Bcd16]"; S7_GenerateENO := "TRUE" } Convert(in := #Temp_9, out => #Temp_9)
      { S7_Templates := "SrcType := Int"; S7_GenerateENO := "TRUE" } Add(in1 := #Temp_9, in2 := 4096, out => #Temp_9)
   END_RUNG
   // the same network as SCL:
   // ENO of a box is taken as its EN; it also drops when the box reports an error
   #Temp_9 := "DB53".Static_15 * 10;
   #Temp_9 := INT_TO_BCD16(#Temp_9);
   #Temp_9 := #Temp_9 + 4096;
END_REGION

REGION Network 15